(* Logix 5000 project; controller PLC_MCC1201_220AP1 vendor 1 type 14 code 164 rev 35.11; software revision 35.00; part 9 of 25 *)
(* tags used below, declared in another part *)
   B3 : DINT[102];
   HMI_Alarm_Reset : BOOL;   // HMI_Alarm_Reset
   HMI_MAN_CMD_WR : UDT_MAN_CMD_WR;
   LEHR_SPEED : ALIAS FOR N60[1];
   M217_M1_DR : AXIS_CIP_DRIVE;
   M218_M1_DR : AXIS_CIP_DRIVE;
   M219_M1_DR : AXIS_CIP_DRIVE;
   M220_M1_DR : AXIS_CIP_DRIVE;
   M2xx_CONVEYOR : MAC_CONVEYOR[20];
   M2xx_CONVEYOR_IN_MOTION : MAC_CONVEYOR_IN_MOTION[20];
   M2xx_CONVEYOR_OUT_MOTION : MAC_CONVEYOR_OUT_MOTION[20];
   TMP_dDirection : DINT;
   TMP_rAcc : REAL;
   TMP_rDec : REAL;
   TMP_rSpeed : REAL;
   TMP_xAlwaysOFF : BOOL;
   TMP_xRun : BOOL;
(* CommandLogic, continued *)

ROUTINE M217_Conveyor_Motion_Output   (* ladder *)
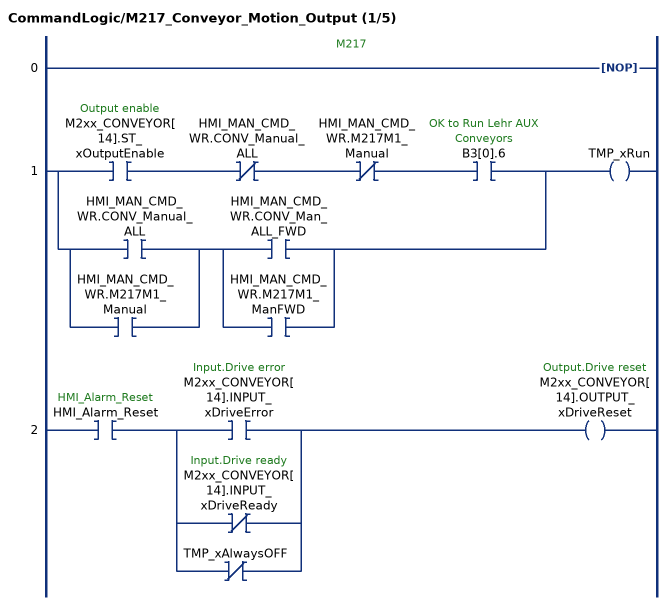
   // M217
   0: NOP();
   1: [XIC(M2xx_CONVEYOR[14].ST_xOutputEnable) XIO(HMI_MAN_CMD_WR.CONV_Manual_ALL) XIO(HMI_MAN_CMD_WR.M217M1_Manual) XIC(B3[0].6) ,[XIC(HMI_MAN_CMD_WR.CONV_Manual_ALL) ,XIC(HMI_MAN_CMD_WR.M217M1_Manual) ] [XIC(HMI_MAN_CMD_WR.CONV_Man_ALL_FWD) ,XIC(HMI_MAN_CMD_WR.M217M1_ManFWD) ] ]OTE(TMP_xRun);
   2: XIC(HMI_Alarm_Reset)[XIC(M2xx_CONVEYOR[14].INPUT_xDriveError) ,XIO(M2xx_CONVEYOR[14].INPUT_xDriveReady) ,XIO(TMP_xAlwaysOFF) ]OTE(M2xx_CONVEYOR[14].OUTPUT_xDriveReset);
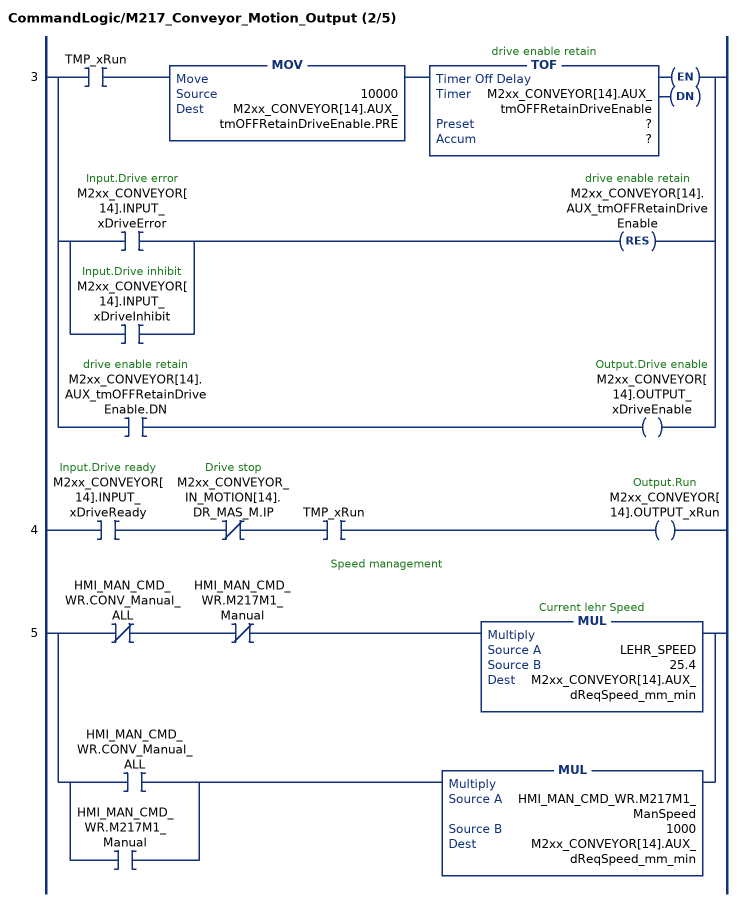
   3: [XIC(TMP_xRun) MOV(10000,M2xx_CONVEYOR[14].AUX_tmOFFRetainDriveEnable.PRE) TOF(M2xx_CONVEYOR[14].AUX_tmOFFRetainDriveEnable,?,?) ,[XIC(M2xx_CONVEYOR[14].INPUT_xDriveError) ,XIC(M2xx_CONVEYOR[14].INPUT_xDriveInhibit) ] RES(M2xx_CONVEYOR[14].AUX_tmOFFRetainDriveEnable) ,XIC(M2xx_CONVEYOR[14].AUX_tmOFFRetainDriveEnable.DN) OTE(M2xx_CONVEYOR[14].OUTPUT_xDriveEnable) ];
   4: XIC(M2xx_CONVEYOR[14].INPUT_xDriveReady)XIO(M2xx_CONVEYOR_IN_MOTION[14].DR_MAS_M.IP)XIC(TMP_xRun)OTE(M2xx_CONVEYOR[14].OUTPUT_xRun);
   // Speed management
   5: [XIO(HMI_MAN_CMD_WR.CONV_Manual_ALL) XIO(HMI_MAN_CMD_WR.M217M1_Manual) MUL(LEHR_SPEED,25.4,M2xx_CONVEYOR[14].AUX_dReqSpeed_mm_min) ,[XIC(HMI_MAN_CMD_WR.CONV_Manual_ALL) ,XIC(HMI_MAN_CMD_WR.M217M1_Manual) ] MUL(HMI_MAN_CMD_WR.M217M1_ManSpeed,1000,M2xx_CONVEYOR[14].AUX_dReqSpeed_mm_min) ];
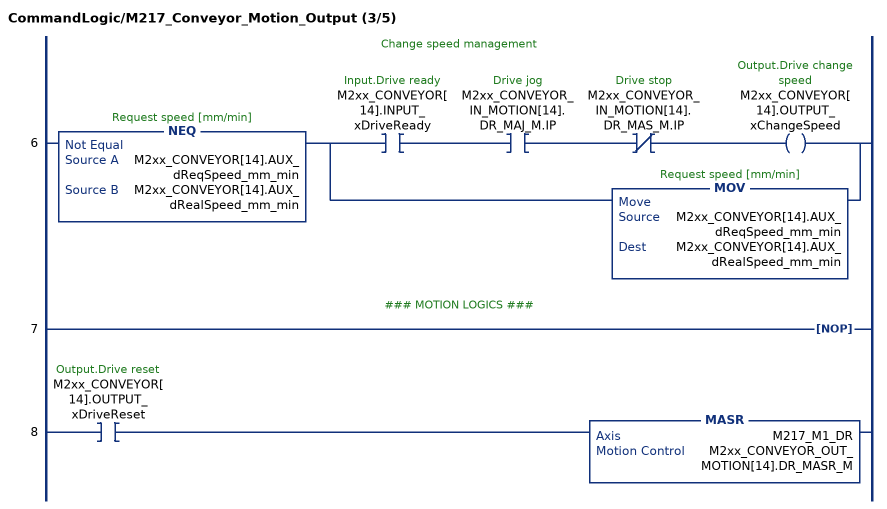
   // Change speed management
   6: NEQ(M2xx_CONVEYOR[14].AUX_dReqSpeed_mm_min,M2xx_CONVEYOR[14].AUX_dRealSpeed_mm_min)[XIC(M2xx_CONVEYOR[14].INPUT_xDriveReady) XIC(M2xx_CONVEYOR_IN_MOTION[14].DR_MAJ_M.IP) XIO(M2xx_CONVEYOR_IN_MOTION[14].DR_MAS_M.IP) OTE(M2xx_CONVEYOR[14].OUTPUT_xChangeSpeed) ,MOV(M2xx_CONVEYOR[14].AUX_dReqSpeed_mm_min,M2xx_CONVEYOR[14].AUX_dRealSpeed_mm_min) ];
   // ### MOTION LOGICS ###
   7: NOP();
   8: XIC(M2xx_CONVEYOR[14].OUTPUT_xDriveReset)MASR(M217_M1_DR,M2xx_CONVEYOR_OUT_MOTION[14].DR_MASR_M);
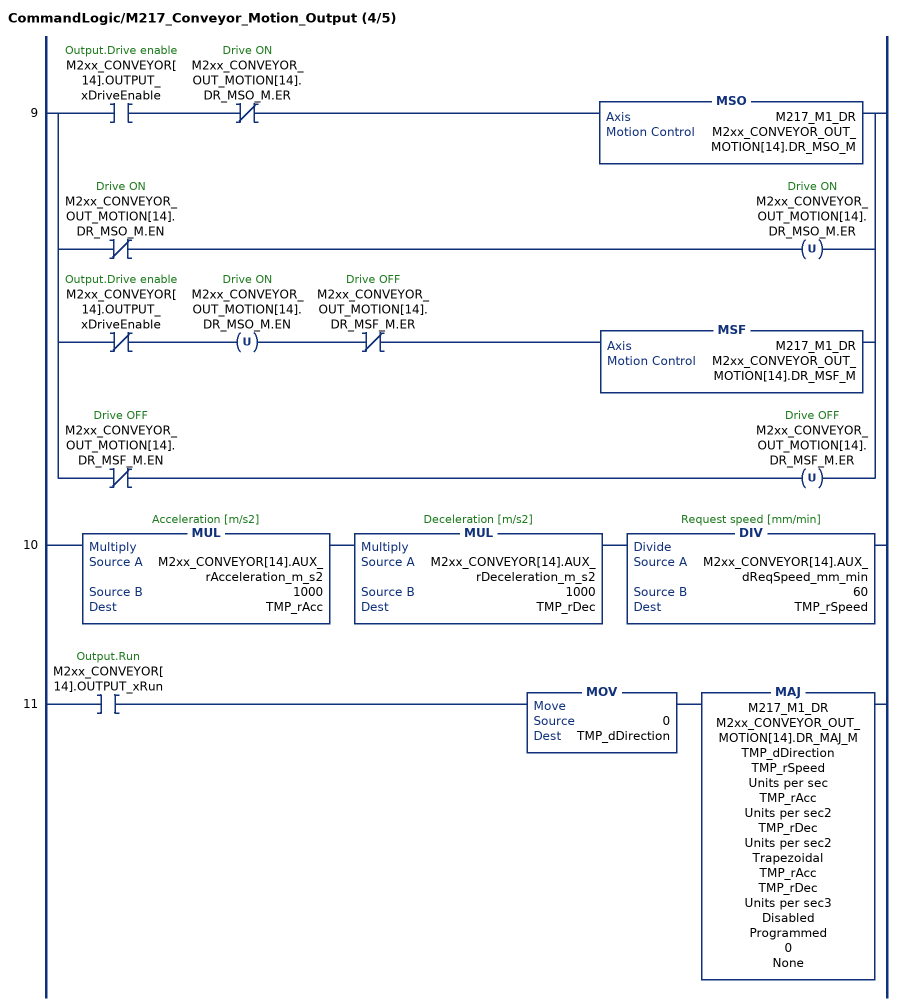
   9: [XIC(M2xx_CONVEYOR[14].OUTPUT_xDriveEnable) XIO(M2xx_CONVEYOR_OUT_MOTION[14].DR_MSO_M.ER) MSO(M217_M1_DR,M2xx_CONVEYOR_OUT_MOTION[14].DR_MSO_M) ,XIO(M2xx_CONVEYOR_OUT_MOTION[14].DR_MSO_M.EN) OTU(M2xx_CONVEYOR_OUT_MOTION[14].DR_MSO_M.ER) ,XIO(M2xx_CONVEYOR[14].OUTPUT_xDriveEnable) OTU(M2xx_CONVEYOR_OUT_MOTION[14].DR_MSO_M.EN) XIO(M2xx_CONVEYOR_OUT_MOTION[14].DR_MSF_M.ER) MSF(M217_M1_DR,M2xx_CONVEYOR_OUT_MOTION[14].DR_MSF_M) ,XIO(M2xx_CONVEYOR_OUT_MOTION[14].DR_MSF_M.EN) OTU(M2xx_CONVEYOR_OUT_MOTION[14].DR_MSF_M.ER) ];
   10: MUL(M2xx_CONVEYOR[14].AUX_rAcceleration_m_s2,1000,TMP_rAcc)MUL(M2xx_CONVEYOR[14].AUX_rDeceleration_m_s2,1000,TMP_rDec)DIV(M2xx_CONVEYOR[14].AUX_dReqSpeed_mm_min,60,TMP_rSpeed);
   11: XIC(M2xx_CONVEYOR[14].OUTPUT_xRun)MOV(0,TMP_dDirection)MAJ(M217_M1_DR,M2xx_CONVEYOR_OUT_MOTION[14].DR_MAJ_M,TMP_dDirection,TMP_rSpeed,Units per sec,TMP_rAcc,Units per sec2,TMP_rDec,Units per sec2,Trapezoidal,TMP_rAcc,TMP_rDec,Units per sec3,Disabled,Programmed,0,None);
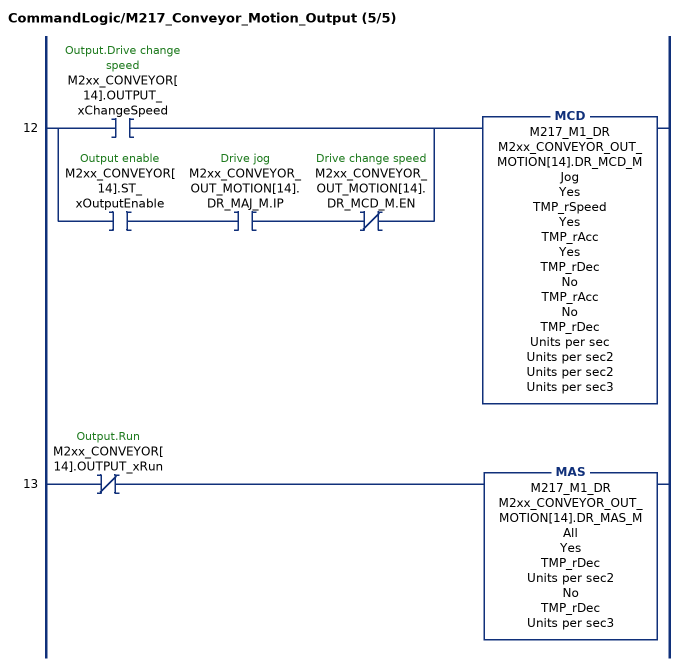
   12: [XIC(M2xx_CONVEYOR[14].OUTPUT_xChangeSpeed) ,XIC(M2xx_CONVEYOR[14].ST_xOutputEnable) XIC(M2xx_CONVEYOR_OUT_MOTION[14].DR_MAJ_M.IP) XIO(M2xx_CONVEYOR_OUT_MOTION[14].DR_MCD_M.EN) ]MCD(M217_M1_DR,M2xx_CONVEYOR_OUT_MOTION[14].DR_MCD_M,Jog,Yes,TMP_rSpeed,Yes,TMP_rAcc,Yes,TMP_rDec,No,TMP_rAcc,No,TMP_rDec,Units per sec,Units per sec2,Units per sec2,Units per sec3);
   13: XIO(M2xx_CONVEYOR[14].OUTPUT_xRun)MAS(M217_M1_DR,M2xx_CONVEYOR_OUT_MOTION[14].DR_MAS_M,All,Yes,TMP_rDec,Units per sec2,No,TMP_rDec,Units per sec3);
END_ROUTINE

ROUTINE M218_Conveyor_Motion_Output   (* ladder *)
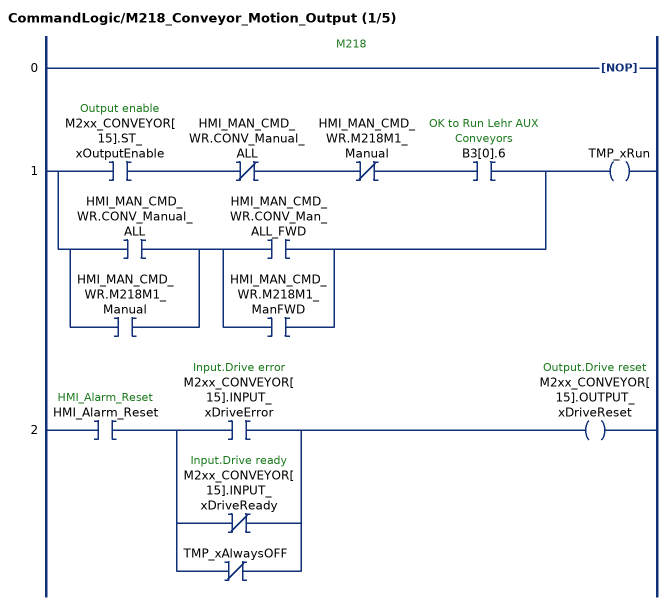
   // M218
   0: NOP();
   1: [XIC(M2xx_CONVEYOR[15].ST_xOutputEnable) XIO(HMI_MAN_CMD_WR.CONV_Manual_ALL) XIO(HMI_MAN_CMD_WR.M218M1_Manual) XIC(B3[0].6) ,[XIC(HMI_MAN_CMD_WR.CONV_Manual_ALL) ,XIC(HMI_MAN_CMD_WR.M218M1_Manual) ] [XIC(HMI_MAN_CMD_WR.CONV_Man_ALL_FWD) ,XIC(HMI_MAN_CMD_WR.M218M1_ManFWD) ] ]OTE(TMP_xRun);
   2: XIC(HMI_Alarm_Reset)[XIC(M2xx_CONVEYOR[15].INPUT_xDriveError) ,XIO(M2xx_CONVEYOR[15].INPUT_xDriveReady) ,XIO(TMP_xAlwaysOFF) ]OTE(M2xx_CONVEYOR[15].OUTPUT_xDriveReset);
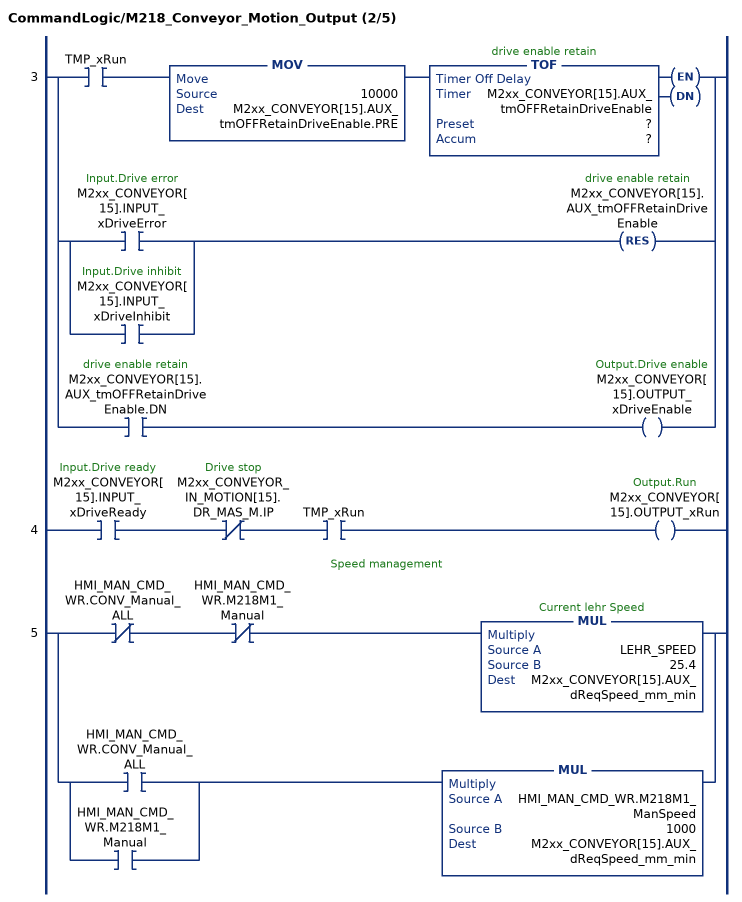
   3: [XIC(TMP_xRun) MOV(10000,M2xx_CONVEYOR[15].AUX_tmOFFRetainDriveEnable.PRE) TOF(M2xx_CONVEYOR[15].AUX_tmOFFRetainDriveEnable,?,?) ,[XIC(M2xx_CONVEYOR[15].INPUT_xDriveError) ,XIC(M2xx_CONVEYOR[15].INPUT_xDriveInhibit) ] RES(M2xx_CONVEYOR[15].AUX_tmOFFRetainDriveEnable) ,XIC(M2xx_CONVEYOR[15].AUX_tmOFFRetainDriveEnable.DN) OTE(M2xx_CONVEYOR[15].OUTPUT_xDriveEnable) ];
   4: XIC(M2xx_CONVEYOR[15].INPUT_xDriveReady)XIO(M2xx_CONVEYOR_IN_MOTION[15].DR_MAS_M.IP)XIC(TMP_xRun)OTE(M2xx_CONVEYOR[15].OUTPUT_xRun);
   // Speed management
   5: [XIO(HMI_MAN_CMD_WR.CONV_Manual_ALL) XIO(HMI_MAN_CMD_WR.M218M1_Manual) MUL(LEHR_SPEED,25.4,M2xx_CONVEYOR[15].AUX_dReqSpeed_mm_min) ,[XIC(HMI_MAN_CMD_WR.CONV_Manual_ALL) ,XIC(HMI_MAN_CMD_WR.M218M1_Manual) ] MUL(HMI_MAN_CMD_WR.M218M1_ManSpeed,1000,M2xx_CONVEYOR[15].AUX_dReqSpeed_mm_min) ];
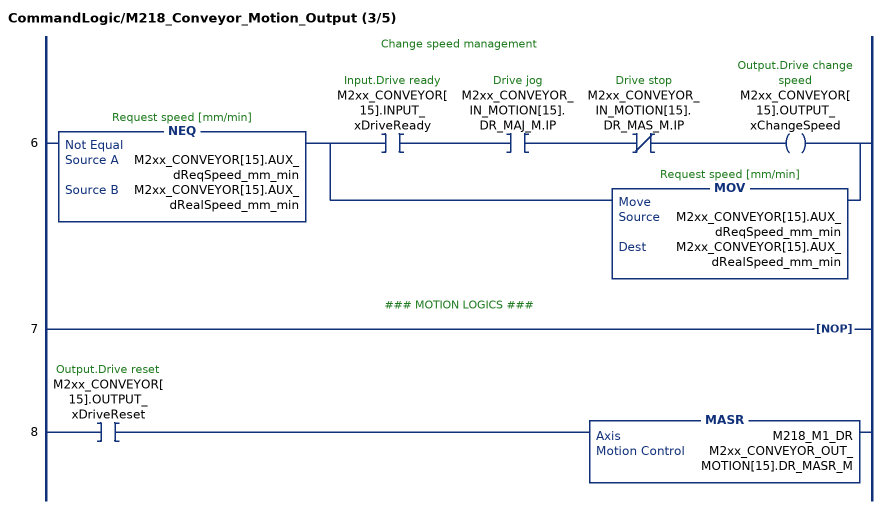
   // Change speed management
   6: NEQ(M2xx_CONVEYOR[15].AUX_dReqSpeed_mm_min,M2xx_CONVEYOR[15].AUX_dRealSpeed_mm_min)[XIC(M2xx_CONVEYOR[15].INPUT_xDriveReady) XIC(M2xx_CONVEYOR_IN_MOTION[15].DR_MAJ_M.IP) XIO(M2xx_CONVEYOR_IN_MOTION[15].DR_MAS_M.IP) OTE(M2xx_CONVEYOR[15].OUTPUT_xChangeSpeed) ,MOV(M2xx_CONVEYOR[15].AUX_dReqSpeed_mm_min,M2xx_CONVEYOR[15].AUX_dRealSpeed_mm_min) ];
   // ### MOTION LOGICS ###
   7: NOP();
   8: XIC(M2xx_CONVEYOR[15].OUTPUT_xDriveReset)MASR(M218_M1_DR,M2xx_CONVEYOR_OUT_MOTION[15].DR_MASR_M);
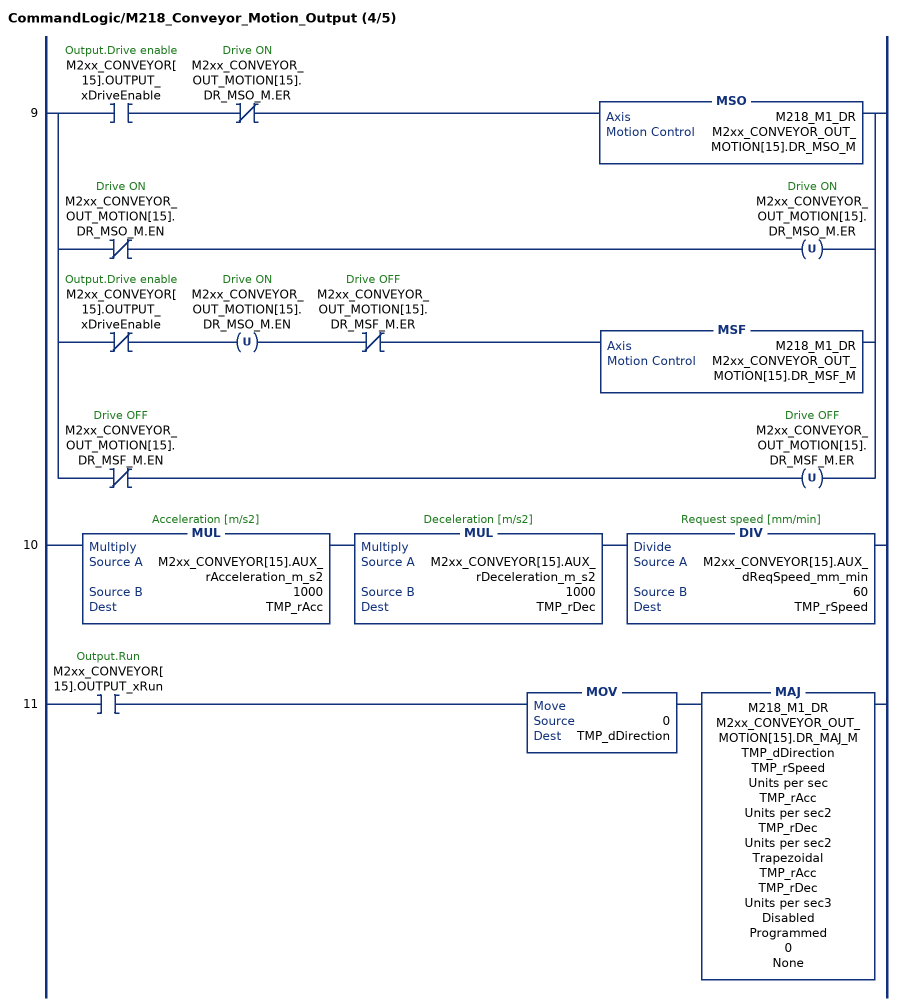
   9: [XIC(M2xx_CONVEYOR[15].OUTPUT_xDriveEnable) XIO(M2xx_CONVEYOR_OUT_MOTION[15].DR_MSO_M.ER) MSO(M218_M1_DR,M2xx_CONVEYOR_OUT_MOTION[15].DR_MSO_M) ,XIO(M2xx_CONVEYOR_OUT_MOTION[15].DR_MSO_M.EN) OTU(M2xx_CONVEYOR_OUT_MOTION[15].DR_MSO_M.ER) ,XIO(M2xx_CONVEYOR[15].OUTPUT_xDriveEnable) OTU(M2xx_CONVEYOR_OUT_MOTION[15].DR_MSO_M.EN) XIO(M2xx_CONVEYOR_OUT_MOTION[15].DR_MSF_M.ER) MSF(M218_M1_DR,M2xx_CONVEYOR_OUT_MOTION[15].DR_MSF_M) ,XIO(M2xx_CONVEYOR_OUT_MOTION[15].DR_MSF_M.EN) OTU(M2xx_CONVEYOR_OUT_MOTION[15].DR_MSF_M.ER) ];
   10: MUL(M2xx_CONVEYOR[15].AUX_rAcceleration_m_s2,1000,TMP_rAcc)MUL(M2xx_CONVEYOR[15].AUX_rDeceleration_m_s2,1000,TMP_rDec)DIV(M2xx_CONVEYOR[15].AUX_dReqSpeed_mm_min,60,TMP_rSpeed);
   11: XIC(M2xx_CONVEYOR[15].OUTPUT_xRun)MOV(0,TMP_dDirection)MAJ(M218_M1_DR,M2xx_CONVEYOR_OUT_MOTION[15].DR_MAJ_M,TMP_dDirection,TMP_rSpeed,Units per sec,TMP_rAcc,Units per sec2,TMP_rDec,Units per sec2,Trapezoidal,TMP_rAcc,TMP_rDec,Units per sec3,Disabled,Programmed,0,None);
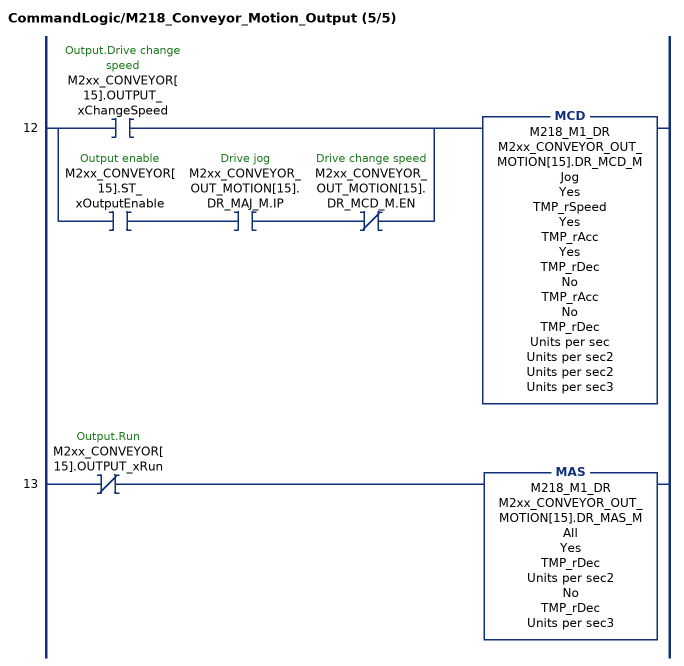
   12: [XIC(M2xx_CONVEYOR[15].OUTPUT_xChangeSpeed) ,XIC(M2xx_CONVEYOR[15].ST_xOutputEnable) XIC(M2xx_CONVEYOR_OUT_MOTION[15].DR_MAJ_M.IP) XIO(M2xx_CONVEYOR_OUT_MOTION[15].DR_MCD_M.EN) ]MCD(M218_M1_DR,M2xx_CONVEYOR_OUT_MOTION[15].DR_MCD_M,Jog,Yes,TMP_rSpeed,Yes,TMP_rAcc,Yes,TMP_rDec,No,TMP_rAcc,No,TMP_rDec,Units per sec,Units per sec2,Units per sec2,Units per sec3);
   13: XIO(M2xx_CONVEYOR[15].OUTPUT_xRun)MAS(M218_M1_DR,M2xx_CONVEYOR_OUT_MOTION[15].DR_MAS_M,All,Yes,TMP_rDec,Units per sec2,No,TMP_rDec,Units per sec3);
END_ROUTINE

ROUTINE M219_Conveyor_Motion_Output   (* ladder *)
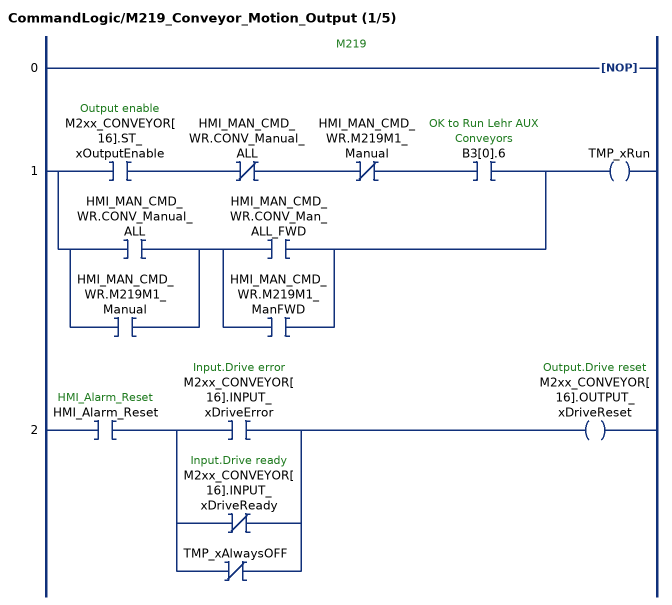
   // M219
   0: NOP();
   1: [XIC(M2xx_CONVEYOR[16].ST_xOutputEnable) XIO(HMI_MAN_CMD_WR.CONV_Manual_ALL) XIO(HMI_MAN_CMD_WR.M219M1_Manual) XIC(B3[0].6) ,[XIC(HMI_MAN_CMD_WR.CONV_Manual_ALL) ,XIC(HMI_MAN_CMD_WR.M219M1_Manual) ] [XIC(HMI_MAN_CMD_WR.CONV_Man_ALL_FWD) ,XIC(HMI_MAN_CMD_WR.M219M1_ManFWD) ] ]OTE(TMP_xRun);
   2: XIC(HMI_Alarm_Reset)[XIC(M2xx_CONVEYOR[16].INPUT_xDriveError) ,XIO(M2xx_CONVEYOR[16].INPUT_xDriveReady) ,XIO(TMP_xAlwaysOFF) ]OTE(M2xx_CONVEYOR[16].OUTPUT_xDriveReset);
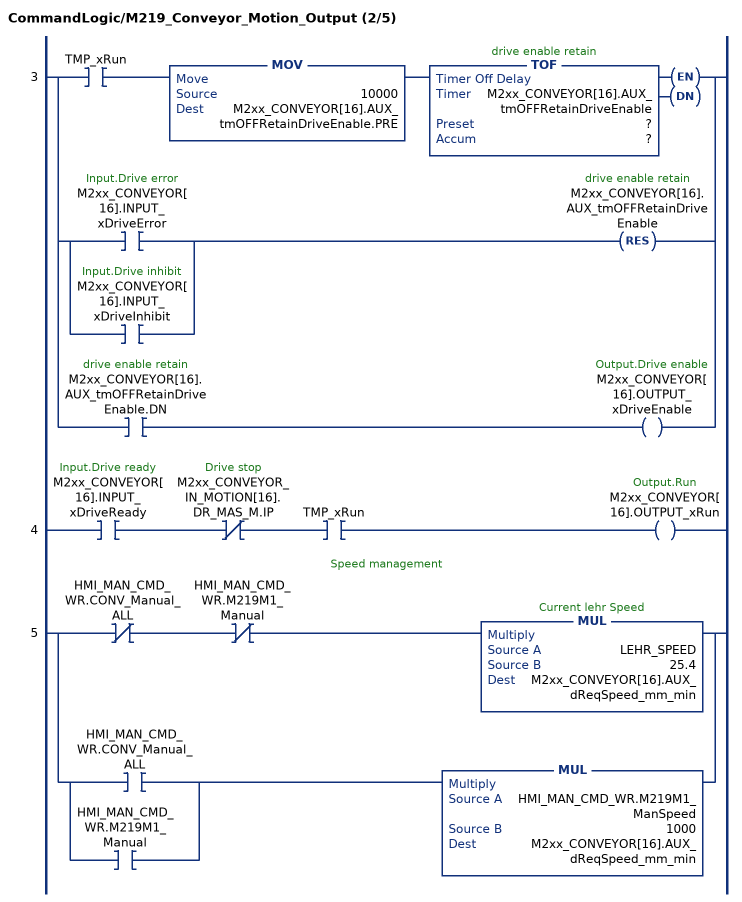
   3: [XIC(TMP_xRun) MOV(10000,M2xx_CONVEYOR[16].AUX_tmOFFRetainDriveEnable.PRE) TOF(M2xx_CONVEYOR[16].AUX_tmOFFRetainDriveEnable,?,?) ,[XIC(M2xx_CONVEYOR[16].INPUT_xDriveError) ,XIC(M2xx_CONVEYOR[16].INPUT_xDriveInhibit) ] RES(M2xx_CONVEYOR[16].AUX_tmOFFRetainDriveEnable) ,XIC(M2xx_CONVEYOR[16].AUX_tmOFFRetainDriveEnable.DN) OTE(M2xx_CONVEYOR[16].OUTPUT_xDriveEnable) ];
   4: XIC(M2xx_CONVEYOR[16].INPUT_xDriveReady)XIO(M2xx_CONVEYOR_IN_MOTION[16].DR_MAS_M.IP)XIC(TMP_xRun)OTE(M2xx_CONVEYOR[16].OUTPUT_xRun);
   // Speed management
   5: [XIO(HMI_MAN_CMD_WR.CONV_Manual_ALL) XIO(HMI_MAN_CMD_WR.M219M1_Manual) MUL(LEHR_SPEED,25.4,M2xx_CONVEYOR[16].AUX_dReqSpeed_mm_min) ,[XIC(HMI_MAN_CMD_WR.CONV_Manual_ALL) ,XIC(HMI_MAN_CMD_WR.M219M1_Manual) ] MUL(HMI_MAN_CMD_WR.M219M1_ManSpeed,1000,M2xx_CONVEYOR[16].AUX_dReqSpeed_mm_min) ];
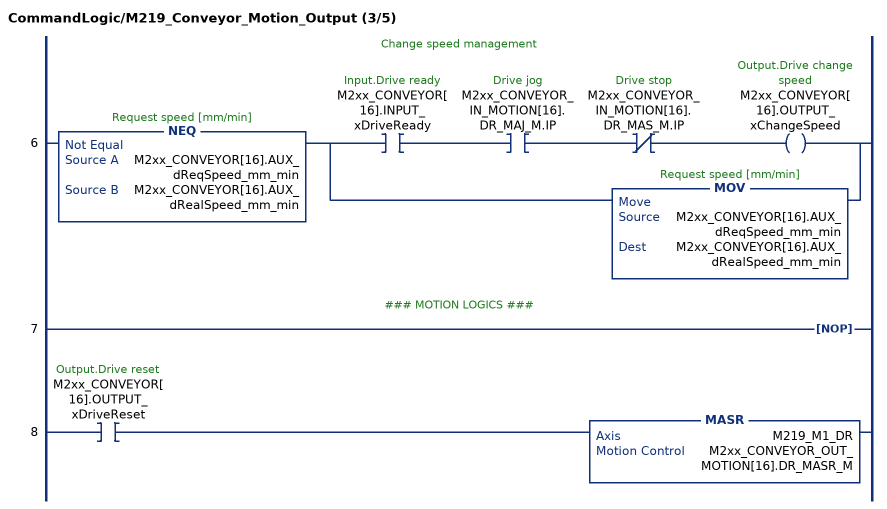
   // Change speed management
   6: NEQ(M2xx_CONVEYOR[16].AUX_dReqSpeed_mm_min,M2xx_CONVEYOR[16].AUX_dRealSpeed_mm_min)[XIC(M2xx_CONVEYOR[16].INPUT_xDriveReady) XIC(M2xx_CONVEYOR_IN_MOTION[16].DR_MAJ_M.IP) XIO(M2xx_CONVEYOR_IN_MOTION[16].DR_MAS_M.IP) OTE(M2xx_CONVEYOR[16].OUTPUT_xChangeSpeed) ,MOV(M2xx_CONVEYOR[16].AUX_dReqSpeed_mm_min,M2xx_CONVEYOR[16].AUX_dRealSpeed_mm_min) ];
   // ### MOTION LOGICS ###
   7: NOP();
   8: XIC(M2xx_CONVEYOR[16].OUTPUT_xDriveReset)MASR(M219_M1_DR,M2xx_CONVEYOR_OUT_MOTION[16].DR_MASR_M);
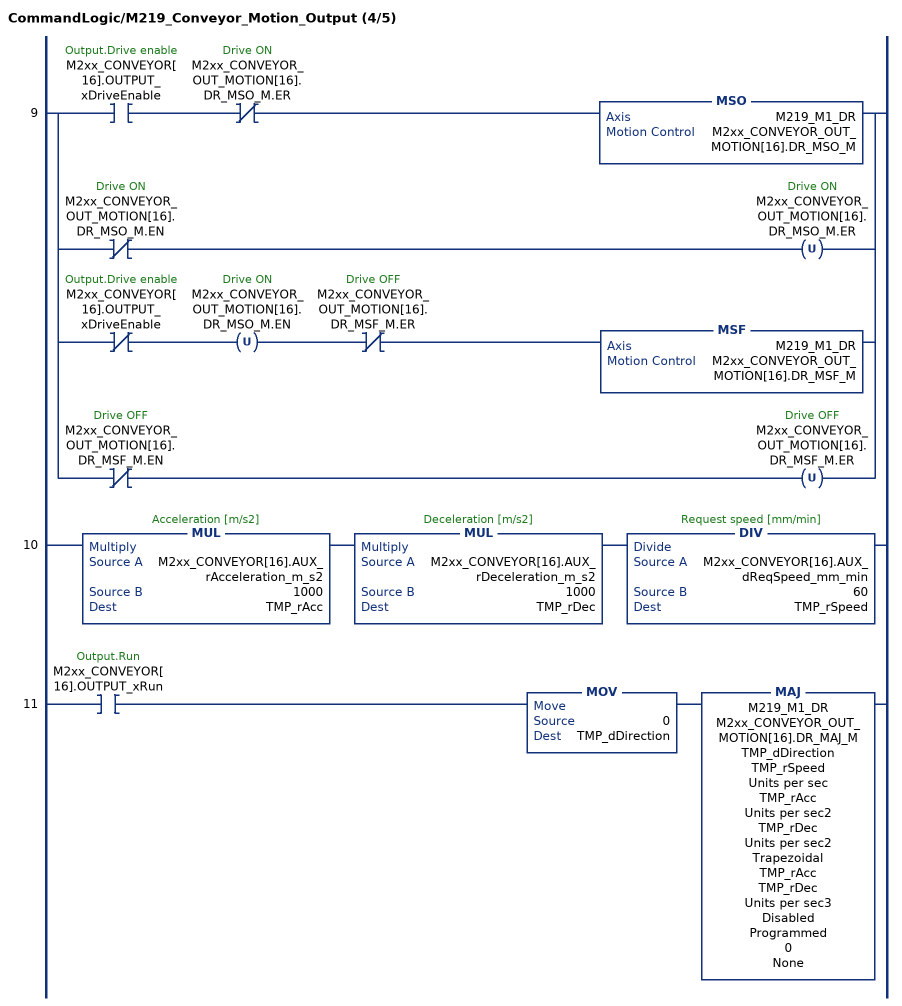
   9: [XIC(M2xx_CONVEYOR[16].OUTPUT_xDriveEnable) XIO(M2xx_CONVEYOR_OUT_MOTION[16].DR_MSO_M.ER) MSO(M219_M1_DR,M2xx_CONVEYOR_OUT_MOTION[16].DR_MSO_M) ,XIO(M2xx_CONVEYOR_OUT_MOTION[16].DR_MSO_M.EN) OTU(M2xx_CONVEYOR_OUT_MOTION[16].DR_MSO_M.ER) ,XIO(M2xx_CONVEYOR[16].OUTPUT_xDriveEnable) OTU(M2xx_CONVEYOR_OUT_MOTION[16].DR_MSO_M.EN) XIO(M2xx_CONVEYOR_OUT_MOTION[16].DR_MSF_M.ER) MSF(M219_M1_DR,M2xx_CONVEYOR_OUT_MOTION[16].DR_MSF_M) ,XIO(M2xx_CONVEYOR_OUT_MOTION[16].DR_MSF_M.EN) OTU(M2xx_CONVEYOR_OUT_MOTION[16].DR_MSF_M.ER) ];
   10: MUL(M2xx_CONVEYOR[16].AUX_rAcceleration_m_s2,1000,TMP_rAcc)MUL(M2xx_CONVEYOR[16].AUX_rDeceleration_m_s2,1000,TMP_rDec)DIV(M2xx_CONVEYOR[16].AUX_dReqSpeed_mm_min,60,TMP_rSpeed);
   11: XIC(M2xx_CONVEYOR[16].OUTPUT_xRun)MOV(0,TMP_dDirection)MAJ(M219_M1_DR,M2xx_CONVEYOR_OUT_MOTION[16].DR_MAJ_M,TMP_dDirection,TMP_rSpeed,Units per sec,TMP_rAcc,Units per sec2,TMP_rDec,Units per sec2,Trapezoidal,TMP_rAcc,TMP_rDec,Units per sec3,Disabled,Programmed,0,None);
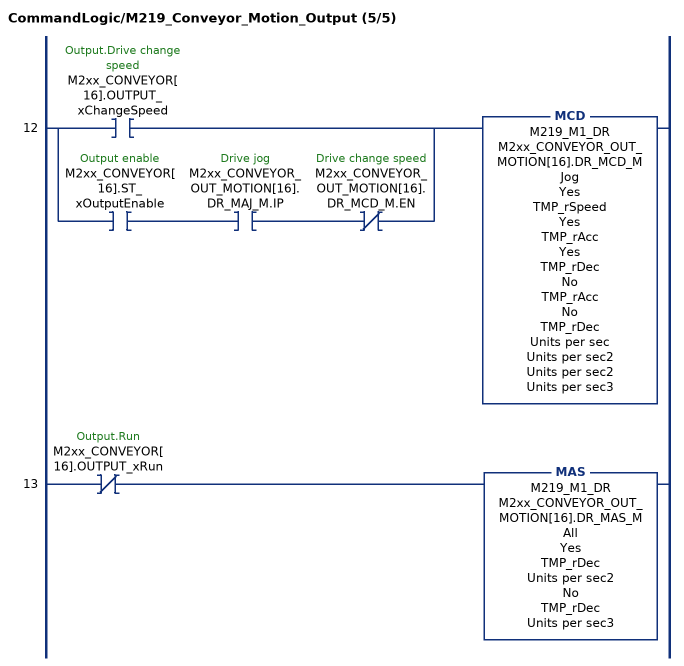
   12: [XIC(M2xx_CONVEYOR[16].OUTPUT_xChangeSpeed) ,XIC(M2xx_CONVEYOR[16].ST_xOutputEnable) XIC(M2xx_CONVEYOR_OUT_MOTION[16].DR_MAJ_M.IP) XIO(M2xx_CONVEYOR_OUT_MOTION[16].DR_MCD_M.EN) ]MCD(M219_M1_DR,M2xx_CONVEYOR_OUT_MOTION[16].DR_MCD_M,Jog,Yes,TMP_rSpeed,Yes,TMP_rAcc,Yes,TMP_rDec,No,TMP_rAcc,No,TMP_rDec,Units per sec,Units per sec2,Units per sec2,Units per sec3);
   13: XIO(M2xx_CONVEYOR[16].OUTPUT_xRun)MAS(M219_M1_DR,M2xx_CONVEYOR_OUT_MOTION[16].DR_MAS_M,All,Yes,TMP_rDec,Units per sec2,No,TMP_rDec,Units per sec3);
END_ROUTINE

ROUTINE M220_Conveyor_Motion_Output   (* ladder *)
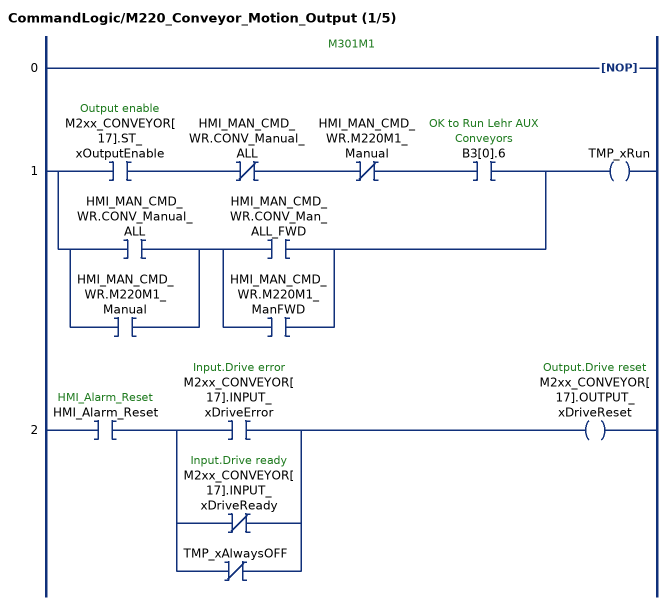
   // M301M1
   0: NOP();
   1: [XIC(M2xx_CONVEYOR[17].ST_xOutputEnable) XIO(HMI_MAN_CMD_WR.CONV_Manual_ALL) XIO(HMI_MAN_CMD_WR.M220M1_Manual) XIC(B3[0].6) ,[XIC(HMI_MAN_CMD_WR.CONV_Manual_ALL) ,XIC(HMI_MAN_CMD_WR.M220M1_Manual) ] [XIC(HMI_MAN_CMD_WR.CONV_Man_ALL_FWD) ,XIC(HMI_MAN_CMD_WR.M220M1_ManFWD) ] ]OTE(TMP_xRun);
   2: XIC(HMI_Alarm_Reset)[XIC(M2xx_CONVEYOR[17].INPUT_xDriveError) ,XIO(M2xx_CONVEYOR[17].INPUT_xDriveReady) ,XIO(TMP_xAlwaysOFF) ]OTE(M2xx_CONVEYOR[17].OUTPUT_xDriveReset);
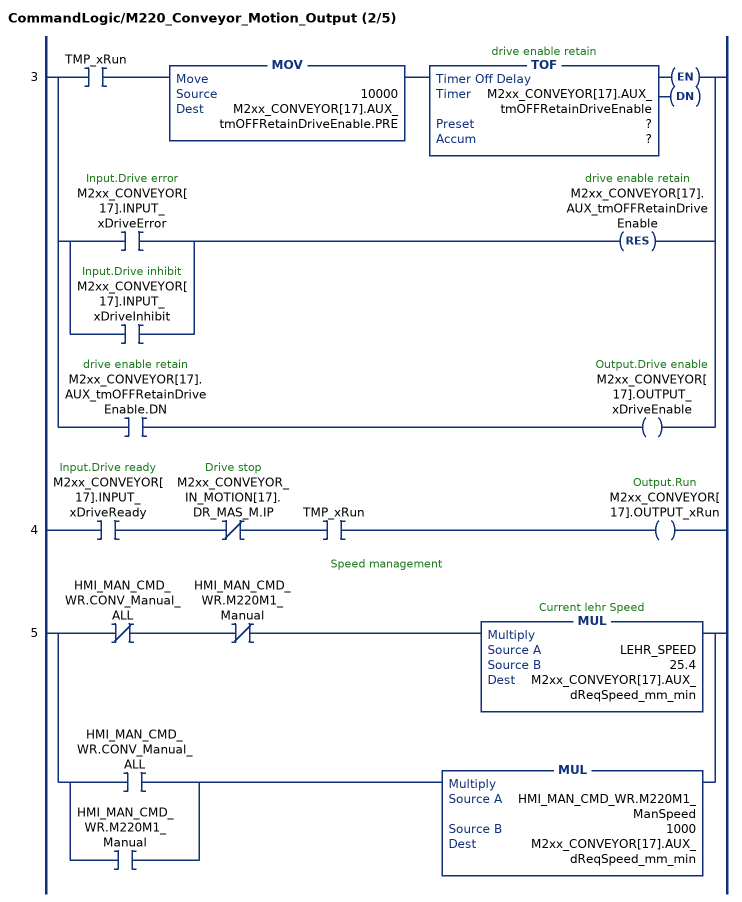
   3: [XIC(TMP_xRun) MOV(10000,M2xx_CONVEYOR[17].AUX_tmOFFRetainDriveEnable.PRE) TOF(M2xx_CONVEYOR[17].AUX_tmOFFRetainDriveEnable,?,?) ,[XIC(M2xx_CONVEYOR[17].INPUT_xDriveError) ,XIC(M2xx_CONVEYOR[17].INPUT_xDriveInhibit) ] RES(M2xx_CONVEYOR[17].AUX_tmOFFRetainDriveEnable) ,XIC(M2xx_CONVEYOR[17].AUX_tmOFFRetainDriveEnable.DN) OTE(M2xx_CONVEYOR[17].OUTPUT_xDriveEnable) ];
   4: XIC(M2xx_CONVEYOR[17].INPUT_xDriveReady)XIO(M2xx_CONVEYOR_IN_MOTION[17].DR_MAS_M.IP)XIC(TMP_xRun)OTE(M2xx_CONVEYOR[17].OUTPUT_xRun);
   // Speed management
   5: [XIO(HMI_MAN_CMD_WR.CONV_Manual_ALL) XIO(HMI_MAN_CMD_WR.M220M1_Manual) MUL(LEHR_SPEED,25.4,M2xx_CONVEYOR[17].AUX_dReqSpeed_mm_min) ,[XIC(HMI_MAN_CMD_WR.CONV_Manual_ALL) ,XIC(HMI_MAN_CMD_WR.M220M1_Manual) ] MUL(HMI_MAN_CMD_WR.M220M1_ManSpeed,1000,M2xx_CONVEYOR[17].AUX_dReqSpeed_mm_min) ];
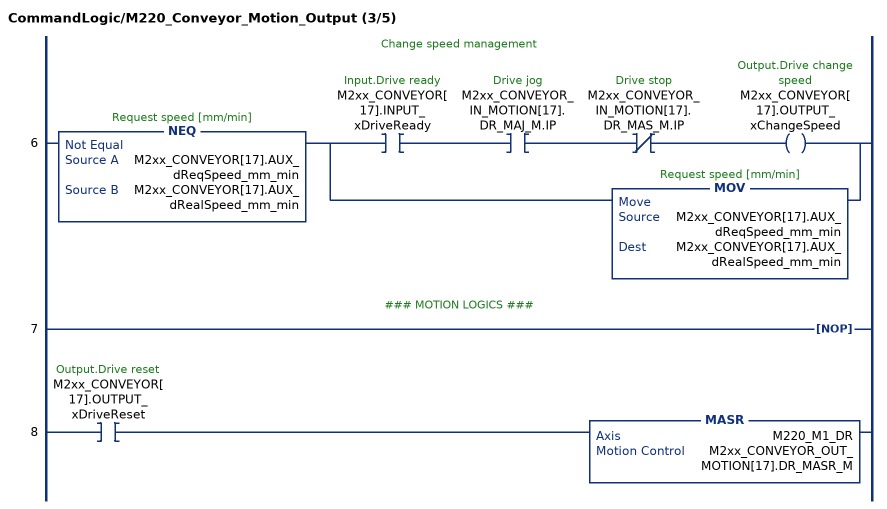
   // Change speed management
   6: NEQ(M2xx_CONVEYOR[17].AUX_dReqSpeed_mm_min,M2xx_CONVEYOR[17].AUX_dRealSpeed_mm_min)[XIC(M2xx_CONVEYOR[17].INPUT_xDriveReady) XIC(M2xx_CONVEYOR_IN_MOTION[17].DR_MAJ_M.IP) XIO(M2xx_CONVEYOR_IN_MOTION[17].DR_MAS_M.IP) OTE(M2xx_CONVEYOR[17].OUTPUT_xChangeSpeed) ,MOV(M2xx_CONVEYOR[17].AUX_dReqSpeed_mm_min,M2xx_CONVEYOR[17].AUX_dRealSpeed_mm_min) ];
   // ### MOTION LOGICS ###
   7: NOP();
   8: XIC(M2xx_CONVEYOR[17].OUTPUT_xDriveReset)MASR(M220_M1_DR,M2xx_CONVEYOR_OUT_MOTION[17].DR_MASR_M);
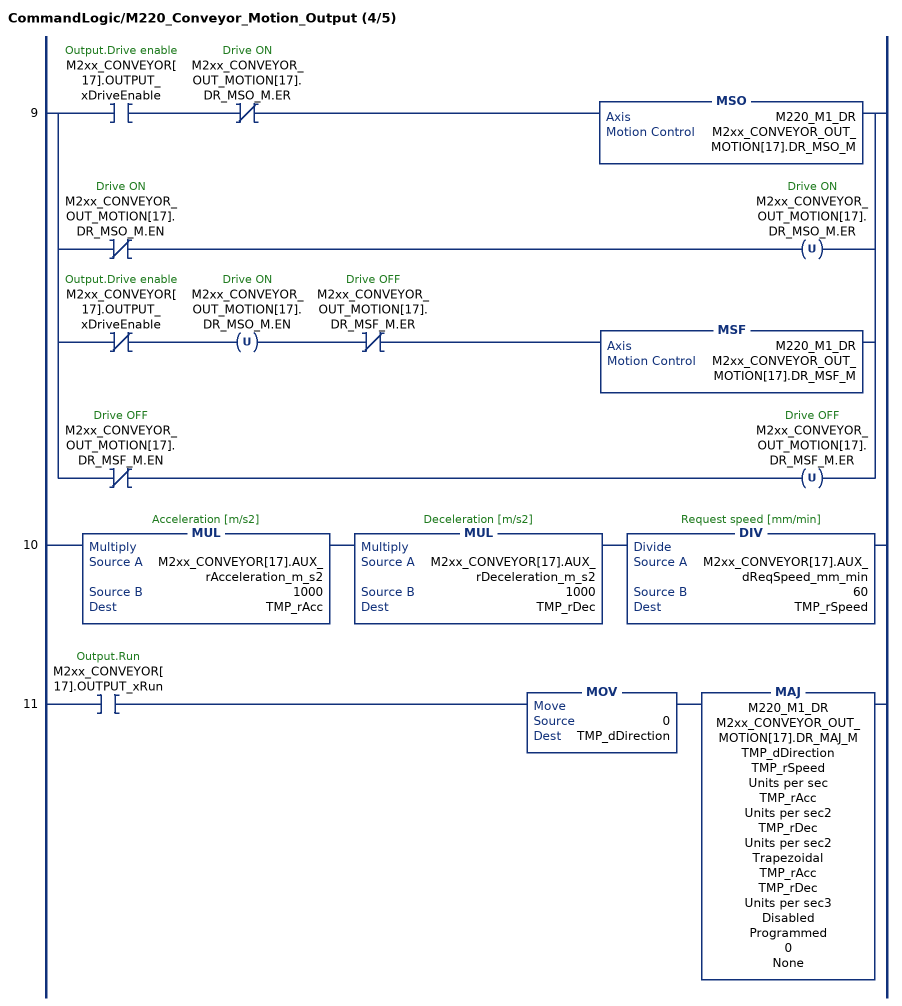
   9: [XIC(M2xx_CONVEYOR[17].OUTPUT_xDriveEnable) XIO(M2xx_CONVEYOR_OUT_MOTION[17].DR_MSO_M.ER) MSO(M220_M1_DR,M2xx_CONVEYOR_OUT_MOTION[17].DR_MSO_M) ,XIO(M2xx_CONVEYOR_OUT_MOTION[17].DR_MSO_M.EN) OTU(M2xx_CONVEYOR_OUT_MOTION[17].DR_MSO_M.ER) ,XIO(M2xx_CONVEYOR[17].OUTPUT_xDriveEnable) OTU(M2xx_CONVEYOR_OUT_MOTION[17].DR_MSO_M.EN) XIO(M2xx_CONVEYOR_OUT_MOTION[17].DR_MSF_M.ER) MSF(M220_M1_DR,M2xx_CONVEYOR_OUT_MOTION[17].DR_MSF_M) ,XIO(M2xx_CONVEYOR_OUT_MOTION[17].DR_MSF_M.EN) OTU(M2xx_CONVEYOR_OUT_MOTION[17].DR_MSF_M.ER) ];
   10: MUL(M2xx_CONVEYOR[17].AUX_rAcceleration_m_s2,1000,TMP_rAcc)MUL(M2xx_CONVEYOR[17].AUX_rDeceleration_m_s2,1000,TMP_rDec)DIV(M2xx_CONVEYOR[17].AUX_dReqSpeed_mm_min,60,TMP_rSpeed);
   11: XIC(M2xx_CONVEYOR[17].OUTPUT_xRun)MOV(0,TMP_dDirection)MAJ(M220_M1_DR,M2xx_CONVEYOR_OUT_MOTION[17].DR_MAJ_M,TMP_dDirection,TMP_rSpeed,Units per sec,TMP_rAcc,Units per sec2,TMP_rDec,Units per sec2,Trapezoidal,TMP_rAcc,TMP_rDec,Units per sec3,Disabled,Programmed,0,None);
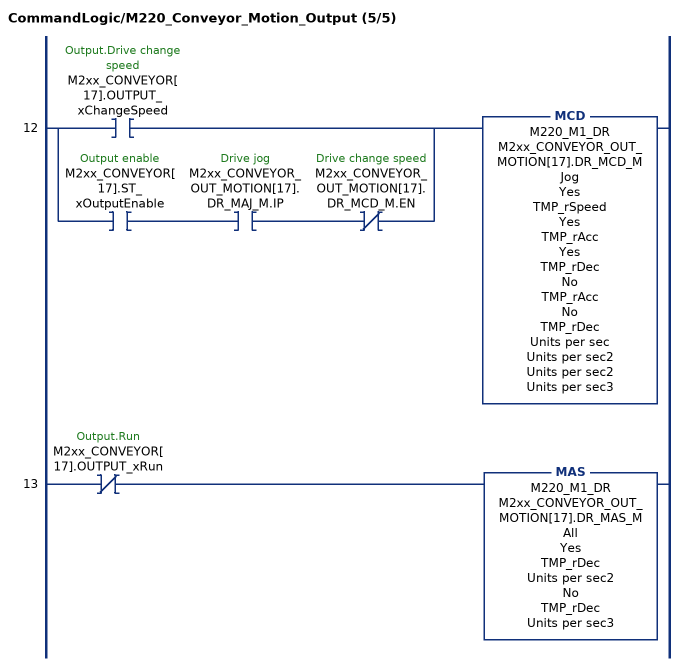
   12: [XIC(M2xx_CONVEYOR[17].OUTPUT_xChangeSpeed) ,XIC(M2xx_CONVEYOR[17].ST_xOutputEnable) XIC(M2xx_CONVEYOR_OUT_MOTION[17].DR_MAJ_M.IP) XIO(M2xx_CONVEYOR_OUT_MOTION[17].DR_MCD_M.EN) ]MCD(M220_M1_DR,M2xx_CONVEYOR_OUT_MOTION[17].DR_MCD_M,Jog,Yes,TMP_rSpeed,Yes,TMP_rAcc,Yes,TMP_rDec,No,TMP_rAcc,No,TMP_rDec,Units per sec,Units per sec2,Units per sec2,Units per sec3);
   13: XIO(M2xx_CONVEYOR[17].OUTPUT_xRun)MAS(M220_M1_DR,M2xx_CONVEYOR_OUT_MOTION[17].DR_MAS_M,All,Yes,TMP_rDec,Units per sec2,No,TMP_rDec,Units per sec3);
END_ROUTINE
